// TIA Portal project "Projekt_Serhii_Bodnia" (V19)
// Vorlageprojekt für das Buch mit Zielsystem S7-1200

(* hardware
DEVICE "S7-1200-Station_1"  S7-1200 Station
   slot 0: "Baugruppenträger_0"  Rack  V1.0
   slot 1: "PLC_1"  CPU 1211C DC/DC/DC  6ES7 211-1AE40-0XB0  V4.1
DEVICE "HMI_1"  KTP900 Basic PN
   slot 0: "HMI_1"  KTP900 Basic PN  6AV2 123-2JB03-0AX0  17.0.0.0
   slot 1: "HMI_RT_1"  KTP900 Basic PN  6AV2 123-2JB03-0AX0  17.0.0.0
   slot 5: "HMI_1.IE_CP_1"  PROFINET Interface  17.0.0.0
      slot 1: "PROFINET Schnittstelle_1"  PROFINET Interface
         slot 1: "Port_1"  Port
*)

// ===== PLC "PLC_1"  CPU 1211C DC/DC/DC =====

VAR_GLOBAL   // PLC tag table "Standard-Variablentabelle"
   "System_Byte" AT %MB10 : Byte;
   "FirstScan" AT %M10.0 : Bool;
   "DiagStatusUpdate" AT %M10.1 : Bool;
   "Clock_Byte" AT %MB0 : Byte;
   "Clock_10Hz" AT %M0.0 : Bool;
   "Clock_5Hz" AT %M0.1 : Bool;
   "Clock_2.5Hz" AT %M0.2 : Bool;
   "Clock_2Hz" AT %M0.3 : Bool;
   "Clock_1.25Hz" AT %M0.4 : Bool;
   "Clock_1Hz" AT %M0.5 : Bool;
   "Clock_0.625Hz" AT %M0.6 : Bool;
   "Clock_0.5Hz" AT %M0.7 : Bool;
END_VAR

VAR_GLOBAL   // PLC tag table "Sensor"
   "Diffuse Sensor 0" AT %I0.0 : Bool;
   "Diffuse Sensor 1" AT %I0.1 : Bool;
   "Diffuse Sensor 2" AT %I0.2 : Bool;
   "Diffuse Sensor 3" AT %I0.3 : Bool;
   "Diffuse Sensor 4" AT %I0.4 : Bool;
   "Diffuse Sensor 5" AT %I0.5 : Bool;
   "Diffuse Sensor 6" AT %I0.6 : Bool;
   "Diffuse Sensor 7" AT %I0.7 : Bool;
   "Diffuse Sensor 8" AT %I1.0 : Bool;
   "Diffuse Sensor 9" AT %I1.1 : Bool;
   "Diffuse Sensor 10" AT %I1.2 : Bool;
   "Diffuse Sensor 11" AT %I1.3 : Bool;
   "Diffuse Sensor 12" AT %I1.4 : Bool;
   "Diffuse Sensor 13" AT %I1.5 : Bool;
   "Diffuse Sensor 14" AT %I1.6 : Bool;
   "Diffuse Sensor 15" AT %I1.7 : Bool;
   "Diffuse Sensor 16" AT %I2.0 : Bool;
   "Diffuse Sensor 17" AT %I2.1 : Bool;
   "Diffuse Sensor 18" AT %I2.2 : Bool;
   "Diffuse Sensor 19" AT %I2.3 : Bool;
   "Diffuse Sensor 20" AT %I2.4 : Bool;
   "Diffuse Sensor 21" AT %I2.5 : Bool;
   "Diffuse Sensor 22" AT %I2.6 : Bool;
   "Diffuse Sensor 23" AT %I2.7 : Bool;
   "Diffuse Sensor 24" AT %I3.0 : Bool;
   "Diffuse Sensor 25" AT %I3.1 : Bool;
   "Diffuse Sensor 26" AT %I3.2 : Bool;
   "Diffuse Sensor 27" AT %I3.3 : Bool;
   "Diffuse Sensor 29" AT %I3.4 : Bool;
   "Emergency Stop 0" AT %I3.6 : Bool;
   "Emergency Stop 1" AT %I3.7 : Bool;
   "Emergency Stop 3" AT %I4.0 : Bool;
   "Left Positioner 1 (Clamped)" AT %I3.5 : Bool;
   "Pick & Place 0 (Box Detected)" AT %I4.1 : Bool;
   "Retroreflective Sensor 1" AT %I4.2 : Bool;
   "Retroreflective Sensor 5" AT %I4.4 : Bool;
   "Retroreflective Sensor 7" AT %I4.5 : Bool;
   "Retroreflective Sensor 10" AT %I4.6 : Bool;
   "Start Button 0" AT %I5.3 : Bool;
   "Start Button 1" AT %I5.0 : Bool;
   "Stop Button 0" AT %I5.1 : Bool;
   "Stop Button 1" AT %I5.2 : Bool;
   "Conveyor Scale 0 Weight (V)" AT %ID30 : Real;
   "Conveyor Scale 1 Weight (V)" AT %ID34 : Real;
   "Tank 1 (Flow Meter)" AT %ID38 : Real;
   "Tank 2 (Flow Meter)" AT %ID42 : Real;
   "Tank 1 (Level Meter)" AT %ID46 : Real;
   "Tank 2 (Level Meter)" AT %ID50 : Real;
   "Vision Sensor 1 (Value)" AT %ID54 : DInt;
   "Retroreflective Sensor 2" AT %I4.3 : Bool;
END_VAR

VAR_GLOBAL   // PLC tag table "Aktor"
   "Belt Conveyor (2m) 0" AT %Q0.0 : Bool;
   "Belt Conveyor (2m) 1" AT %Q0.1 : Bool;
   "Belt Conveyor (2m) 2" AT %Q0.2 : Bool;
   "Belt Conveyor (2m) 3" AT %Q0.3 : Bool;
   "Belt Conveyor (2m) 4" AT %Q0.4 : Bool;
   "Belt Conveyor (4m) 0" AT %Q0.7 : Bool;
   "Belt Conveyor (4m) 2" AT %Q1.0 : Bool;
   "Belt Conveyor (4m) 3" AT %Q1.1 : Bool;
   "Belt Conveyor (4m) 5" AT %Q1.2 : Bool;
   "Belt Conveyor (4m) 6" AT %Q1.3 : Bool;
   "Belt Conveyor (4m) 7" AT %Q1.4 : Bool;
   "Belt Conveyor (6m) 2" AT %Q1.5 : Bool;
   "Belt Conveyor (2m) 6" AT %Q0.5 : Bool;
   "Belt Conveyor (2m) 7" AT %Q0.6 : Bool;
   "Conveyor Scale 0 (+)" AT %Q1.6 : Bool;
   "Conveyor Scale 1 (+)" AT %Q1.7 : Bool;
   "Curved Belt Conveyor 1 CW" AT %Q2.0 : Bool;
   "Curved Belt Conveyor 0 CCW" AT %Q2.1 : Bool;
   "Left Positioner 1 (Clamp)" AT %Q2.2 : Bool;
   "Emitter 1 (Emit)" AT %Q2.3 : Bool;
   "Emitter 3 (Emit)" AT %Q2.4 : Bool;
   "Emitter 4 (Emit)" AT %Q2.5 : Bool;
   "Remover 0 (Remove)" AT %Q2.6 : Bool;
   "Remover 1 (Remove)" AT %Q2.7 : Bool;
   "Remover 2 (Remove)" AT %Q3.0 : Bool;
   "Remover 3 (Remove)" AT %Q3.1 : Bool;
   "Roller Conveyor (2m) 0" AT %Q3.2 : Bool;
   "Roller Conveyor (2m) 1" AT %Q3.3 : Bool;
   "Roller Conveyor (2m) 3" AT %Q3.4 : Bool;
   "Roller Conveyor (4m) 0" AT %Q3.5 : Bool;
   "Pusher 0" AT %Q3.6 : Bool;
   "Pusher 3" AT %Q3.7 : Bool;
   "Pivot Arm Sorter 0 Turn" AT %Q4.0 : Bool;
   "Pivot Arm Sorter 0 Belt (+)" AT %Q4.1 : Bool;
   "Pick & Place 0 (Grab)" AT %Q4.2 : Bool;
   "Start Button 0 (Light)" AT %Q4.3 : Bool;
   "Start Button 1 (Light)" AT %Q4.4 : Bool;
   "Stop Button 0 (Light)" AT %Q4.5 : Bool;
   "Stop Button 1 (Light)" AT %Q4.6 : Bool;
   "Stack Light 0 (Green)" AT %Q4.7 : Bool;
   "Stack Light 0 (Red)" AT %Q5.0 : Bool;
   "Stack Light 0 (Yellow)" AT %Q5.1 : Bool;
   "Stack Light 1 (Green)" AT %Q5.2 : Bool;
   "Stack Light 1 (Red)" AT %Q5.3 : Bool;
   "Stack Light 1 (Yellow)" AT %Q5.4 : Bool;
   "Warning Light 1" AT %Q5.5 : Bool;
   "Pick & Place 0  X Set Point (V)" AT %QD34 : Real;
   "Pick & Place 0  Y Set Point (V)" AT %QD30 : Real;
   "Pick & Place 0  Z Set Point (V)" AT %QD38 : Real;
   "Tank 1 (Fill Valve)" AT %QD46 : Real;
   "Tank 2 (Fill Valve)" AT %QD50 : Real;
   "Tank 1 (Discharge Valve)" AT %QD54 : Real;
   "Tank 2 (Discharge Valve)" AT %QD58 : Real;
END_VAR

VAR_GLOBAL   // PLC tag table "Merker"
   "FlOp_P_Activate" AT %I4.7 : Bool;
END_VAR

TYPE "Getränk"
   STRUCT
      Tankfüllvolumen : Real;
      Dosiervolumen : Real;
      VAR_Rezeptur : Int;
      VAR_Rezeptur_Datensatz : Int;
   END_STRUCT;
END_TYPE

DATA_BLOCK "FB_Laufzeit_DB"   // DB1
{ S7_Optimized_Access := 'TRUE' }
VERSION : 0.1
// stored: InstanceOfName FB_Laufzeit
"FB_Laufzeit"
BEGIN
END_DATA_BLOCK

DATA_BLOCK "FB_Transport_Band_DB_1"   // DB2
{ S7_Optimized_Access := 'TRUE' }
VERSION : 0.1
// stored: InstanceOfName FB_Transport_Band
"FB_Transport_Band"
BEGIN
END_DATA_BLOCK

DATA_BLOCK "GDB_PLC"   // DB3
{ S7_Optimized_Access := 'TRUE' }
VERSION : 0.1
   VAR
      Dosierung_Start_Linie_0 : Bool;
      Dosierung_Start_Linie_1 : Bool;
      Dosing_Activate_Linie_0 : Bool;
      Dosing_Activate_Linie_1 : Bool;
      Eingabe_Level_norm_Linie_0 : Real;
      Eingabe_Level_norm_Linie_1 : Real;
      Tank_0_Level_norm : Real;
      Tank_1_Level_norm : Real;
      Start_Modus_Hauptleitung : Bool;
      Start_Modus_Linie_0 : Bool;
      Licht_in_Betrieb : Bool;
      Licht_außer_Betrieb : Bool;
      Licht_Alarm : Bool;
      Start_Modus_Linie_1 : Bool;
      Stop_Modus_Hauptleitung : Bool;
      Stop_Modus_Linie_0 : Bool;
      Stop_Modus_Linie_1 : Bool;
      Not_Aus_Modus : Bool;
      Füllventil_closed_Linie_0 : Bool;
      Füllventil_closed_Linie_1 : Bool;
      Altuell_Gewicht_Linie_0 : Real;
      Altuell_Gewicht_Linie_1 : Real;
      Gesamtteile_Linie_0 : Int;
      Gesamtteile_Linie_1 : Int;
      Ausschuss_Linie_0 : Int;
      Ausschuss_Linie_1 : Int;
      Anzahl_Paletten : Int;
      Anzahl_Kanister_Packungbereich : Int;
      Anzahl_Kanister_Tr_Band_Halle_2 : Int;
      Tankfüllvolumen_0 : Real;
      Tankfüllvolumen_1 : Real;
      Dosiervolumen_0 : Real;
      Dosiervolumen_1 : Real;
      Ready_to_Send_Teil_Band_Linie_3_0 : Bool;
      Acknowledge_Teil_Greifen_Linie_0 : Bool;
      Palette_voll_Linie_0 : Bool;
      Palette_voll_Linie_1 : Bool;
      Ready_To_Receive_Teil_Palette_Linie_0 : Bool;
      Ready_To_Receive_Teil_Palette_Linie_1 : Bool;
      Ready_To_Send_Teil_Wage_Linie_0 : Bool;
      Ready_To_Send_Teil_Band_2_Linie_0 : Bool;
      Ready_to_Receive_Teil_Band_3_Linie_0 : Bool;
      Run_Hours : Int;
      Run_Minutes : Int;
      Run_Seconds : Int;
      Störung : Array[0..16] of Bool;
   END_VAR
BEGIN
END_DATA_BLOCK

DATA_BLOCK "FB_Tank_DB"   // DB4
{ S7_Optimized_Access := 'TRUE' }
VERSION : 0.1
// stored: InstanceOfName FB_Tank
"FB_Tank"
BEGIN
END_DATA_BLOCK

DATA_BLOCK "FB_Dose_Control_DB"   // DB5
{ S7_Optimized_Access := 'TRUE' }
VERSION : 0.1
// stored: InstanceOfName FB_Dose_Control
"FB_Dose_Control"
BEGIN
END_DATA_BLOCK

DATA_BLOCK "GDB_HMI"   // DB6
{ S7_Optimized_Access := 'TRUE' }
VERSION : 0.1
   VAR
      Meldung_HMI : Int;
      Quittierung_HMI : Int;
      Tankfüllvolumen_HMI : Int;
      Dosiervolumen_HMI : Int;
      Füllmenge_Linie_0 : Real;
      Füllmenge_Linie_1 : Real;
      Reset_Gesamtteile_0 : Bool;
      Reset_Gesamtteile_1 : Bool;
      Reset_Ausschluss_0 : Bool;
      Reset_Ausschluss_1 : Bool;
      NotAus_HMI : Bool;
      Haupt_Stop_HMI : Bool;
   END_VAR
BEGIN
END_DATA_BLOCK

DATA_BLOCK "GDB_Getränk"   // DB7
{ S7_Optimized_Access := 'TRUE' }
VERSION : 0.1
   VAR
      Getränk_Linie_0 : "Getränk";
      Getränk_Linie_1 : "Getränk";
   END_VAR
BEGIN
END_DATA_BLOCK

DATA_BLOCK "FB_Transport_Band_DB_2"   // DB8
{ S7_Optimized_Access := 'TRUE' }
VERSION : 0.1
// stored: InstanceOfName FB_Transport_Band
"FB_Transport_Band"
BEGIN
END_DATA_BLOCK

DATA_BLOCK "FB_Mode_Manager_DB"   // DB9
{ S7_Optimized_Access := 'TRUE' }
VERSION : 0.1
// stored: InstanceOfName FB_Mode_Manager
"FB_Mode_Manager"
BEGIN
END_DATA_BLOCK

DATA_BLOCK "FB_Transport_Band_DB"   // DB10
{ S7_Optimized_Access := 'TRUE' }
VERSION : 0.1
// stored: InstanceOfName FB_Transport_Band
"FB_Transport_Band"
BEGIN
END_DATA_BLOCK

DATA_BLOCK "FB_AbfüllmaschineBand_SCL_DB"   // DB11
{ S7_Optimized_Access := 'TRUE' }
VERSION : 0.1
// stored: InstanceOfName FB_AbfüllmaschineBand_SCL
"FB_AbfüllmaschineBand_SCL"
BEGIN
END_DATA_BLOCK

DATA_BLOCK "FB_Gewichtkontrolle_SCL_DB"   // DB12
{ S7_Optimized_Access := 'TRUE' }
VERSION : 0.1
// stored: InstanceOfName FB_Gewichtkontrolle_SCL
"FB_Gewichtkontrolle_SCL"
BEGIN
END_DATA_BLOCK

DATA_BLOCK "FB_Transport_Band_DB_3"   // DB13
{ S7_Optimized_Access := 'TRUE' }
VERSION : 0.1
// stored: InstanceOfName FB_Transport_Band
"FB_Transport_Band"
BEGIN
END_DATA_BLOCK

DATA_BLOCK "FB_Sortierabschnitt_DB"   // DB14
{ S7_Optimized_Access := 'TRUE' }
VERSION : 0.1
// stored: InstanceOfName FB_Sortierabschnitt
"FB_Sortierabschnitt"
BEGIN
END_DATA_BLOCK

DATA_BLOCK "FB_Transport_Band_DB_4"   // DB15
{ S7_Optimized_Access := 'TRUE' }
VERSION : 0.1
// stored: InstanceOfName FB_Transport_Band
"FB_Transport_Band"
BEGIN
END_DATA_BLOCK

DATA_BLOCK "FB_Band mit Positionierleisten_DB"   // DB16
{ S7_Optimized_Access := 'TRUE' }
VERSION : 0.1
// stored: InstanceOfName FB_Band mit Positionierleisten
"FB_Band mit Positionierleisten"
BEGIN
END_DATA_BLOCK

DATA_BLOCK "FB_Palette_Linie_0_DB"   // DB17
{ S7_Optimized_Access := 'TRUE' }
VERSION : 0.1
// stored: InstanceOfName FB_Palette_Linie
"FB_Palette_Linie"
BEGIN
END_DATA_BLOCK

DATA_BLOCK "FB_Pick & Place_DB"   // DB18
{ S7_Optimized_Access := 'TRUE' }
VERSION : 0.1
// stored: InstanceOfName FB_Pick & Place
"FB_Pick & Place"
BEGIN
END_DATA_BLOCK

DATA_BLOCK "FB_Tank_DB_1"   // DB19
{ S7_Optimized_Access := 'TRUE' }
VERSION : 0.1
// stored: InstanceOfName FB_Tank
"FB_Tank"
BEGIN
END_DATA_BLOCK

DATA_BLOCK "FB_AbfüllmaschineBand_SCL_DB_1"   // DB20
{ S7_Optimized_Access := 'TRUE' }
VERSION : 0.1
// stored: InstanceOfName FB_AbfüllmaschineBand_SCL
"FB_AbfüllmaschineBand_SCL"
BEGIN
END_DATA_BLOCK

DATA_BLOCK "FB_Dose_Control_DB_1"   // DB21
{ S7_Optimized_Access := 'TRUE' }
VERSION : 0.1
// stored: InstanceOfName FB_Dose_Control
"FB_Dose_Control"
BEGIN
END_DATA_BLOCK

DATA_BLOCK "FB_Gewichtkontrolle_SCL_DB_1"   // DB22
{ S7_Optimized_Access := 'TRUE' }
VERSION : 0.1
// stored: InstanceOfName FB_Gewichtkontrolle_SCL
"FB_Gewichtkontrolle_SCL"
BEGIN
END_DATA_BLOCK

DATA_BLOCK "FB_Transport_Band_DB_5"   // DB23
{ S7_Optimized_Access := 'TRUE' }
VERSION : 0.1
// stored: InstanceOfName FB_Transport_Band
"FB_Transport_Band"
BEGIN
END_DATA_BLOCK

DATA_BLOCK "FB_Transport_Band_DB_6"   // DB24
{ S7_Optimized_Access := 'TRUE' }
VERSION : 0.1
// stored: InstanceOfName FB_Transport_Band
"FB_Transport_Band"
BEGIN
END_DATA_BLOCK

DATA_BLOCK "FB_Transport_Band_DB_7"   // DB25
{ S7_Optimized_Access := 'TRUE' }
VERSION : 0.1
// stored: InstanceOfName FB_Transport_Band
"FB_Transport_Band"
BEGIN
END_DATA_BLOCK

DATA_BLOCK "FB_Transportbad mit Verzögerung_DB"   // DB26
{ S7_Optimized_Access := 'TRUE' }
VERSION : 0.1
// stored: InstanceOfName FB_Transportbad mit Verzögerung
"FB_Transportbad mit Verzögerung"
BEGIN
END_DATA_BLOCK

DATA_BLOCK "FB_Transport_T-Band_DB"   // DB27
{ S7_Optimized_Access := 'TRUE' }
VERSION : 0.1
// stored: InstanceOfName FB_Transport_T-Band
"FB_Transport_T-Band"
BEGIN
END_DATA_BLOCK

DATA_BLOCK "FB_Transportbad mit Verzögerung_DB_1"   // DB28
{ S7_Optimized_Access := 'TRUE' }
VERSION : 0.1
// stored: InstanceOfName FB_Transportbad mit Verzögerung
"FB_Transportbad mit Verzögerung"
BEGIN
END_DATA_BLOCK

FUNCTION_BLOCK "FB_Gewichtkontrolle_SCL"   // FB1, SCL
{ S7_Optimized_Access := 'TRUE' }
VERSION : 0.1
   VAR_INPUT
      Start_Mode : Bool;
      Stop_Mode : Bool;
      NotAus_Mode : Bool;
      LS_Einlauf : Bool;
      LS_Mitte : Bool;
      LS_Auslauf : Bool;
      LS_Wage : Bool;
      LS_Pusher : Bool;
      Gewichtsskala : Real;
      Referenz_Gewicht : Real;
      Reset_CTU_Gesamtteile : Bool;
      Reset_CTU_Ausschuss : Bool;
      Quittierung : Bool;
   END_VAR
   VAR_OUTPUT
      Wage_Band : Bool;
      Pusher_Band : Bool;
      Gewicht_Kg : Real;
      Remoover : Bool;
      Pusher : Bool;
      Out_Gesamtteile : Int;
      Out_Ausschuss : Int;
      Ready_To_Send_Teil : Bool;
      Störung : Bool;
   END_VAR
   VAR
      iSchritt : Int;
      Trigger_Pos_LS_Einlauf : R_TRIG;
      Trigger_Neg_LS_Auslauf : F_TRIG;
      Trigger_Pos_LS_Mitte : R_TRIG;
      Trigger_Neg_LS_Mitte : F_TRIG;
      Trigger_Neg_LS_Wage : F_TRIG;
      Trigger_Neg_LS_Pusher : F_TRIG;
      TON_weit_Wiegung_1000ms : TON_TIME;
      TON_Puscher_100ms : TON_TIME;
      TON_Ende_weit_1000ms : TON_TIME;
      TOF_2000ms : TOF_TIME;
      Actuell_Gewicht : Real;
      Gewicht_Norm : Real;
      Speichen_Gewicht : Real;
      Gesamtteile : Int;
      Ausschuss : Int;
      TON_Störung_LS_Wage : TON_TIME;
      TON_Störung_LS_Mitte : TON_TIME;
      TON_Störung_LS_Pusher : TON_TIME;
      TON_Störung_Auslauf : TON_TIME;
      M_Störung : Bool;
      M_Wage_Band : Bool;
      M_Pusher_Band : Bool;
   END_VAR
   VAR CONSTANT
      Toleranz : Real := 1.02;
   END_VAR
BEGIN
   REGION NotAus & Störung
       IF #NotAus_Mode OR #M_Störung THEN
           // Bei Not-Aus or Störung sofortiger Rücksprung in den Initialschritt (Schritt 0)
           #iSchritt := 0;
       END_IF;
   END_REGION

   REGION Reset
       IF #Reset_CTU_Gesamtteile OR #NotAus_Mode OR "FirstScan" THEN
           // Gesamtteilezähler zurücksetzen: bei HMI-Anforderung, Not-Aus oder Erstaufruf
           #Gesamtteile := 0;
       END_IF;

       IF #Reset_CTU_Ausschuss OR #NotAus_Mode OR "FirstScan" THEN
           // Ausschusszähler zurücksetzen: bei HMI-Anforderung, Not-Aus oder Erstaufruf
           #Ausschuss := 0;

       END_IF;

   END_REGION

   REGION Flankenabfragen
       #Trigger_Pos_LS_Einlauf(CLK := #LS_Einlauf); 
       #Trigger_Pos_LS_Mitte(CLK := #LS_Mitte);     
       #Trigger_Neg_LS_Mitte(CLK := #LS_Mitte);
       #Trigger_Neg_LS_Auslauf(CLK := #LS_Auslauf);
       #Trigger_Neg_LS_Wage(CLK := #LS_Wage);
       #Trigger_Neg_LS_Pusher(CLK := #LS_Pusher);
   END_REGION

   REGION Timers
       // Wiegezeit: 500ms Wartezeit für stabile Gewichtsmessung (Schritt 2)
       #TON_weit_Wiegung_1000ms(IN := (#iSchritt = 2),
                                PT := T#500ms);
       // Pusher-Impuls: 100ms Aktivierungszeit für Pusher-Zylinder (Schritt 11)
       #TON_Puscher_100ms(IN := #iSchritt = 11,
                          PT := T#100ms);
       // Remover-Wartezeit: 1000ms bis Remover das Ausschussteil aufgenommen hat (Schritt 12)
       #TON_Ende_weit_1000ms(IN := (#iSchritt = 12),
                             PT := T#1000ms);
       // Anzeigedauer Gewicht: Messwert 2 Sekunden nach Wiegung sichtbar halten (Schritt 2)
       #TOF_2000ms(IN := (#iSchritt = 2),
                   PT := T#2000ms);
       // Störungserkennung: wenn Licht_Sensors länger als 10s aktiv und Band läuft → Stau

       #TON_Störung_LS_Wage(IN := #LS_Wage AND #M_Wage_Band AND NOT #Stop_Mode,
                            PT := T#10s);
       #TON_Störung_LS_Mitte(IN := #LS_Mitte AND #M_Wage_Band AND NOT #Stop_Mode,
                             PT := T#10s);
       #TON_Störung_LS_Pusher(IN := #LS_Pusher AND #M_Pusher_Band AND NOT #Stop_Mode,
                             PT := T#10s);
       #TON_Störung_Auslauf(IN := #LS_Auslauf AND #M_Pusher_Band AND NOT #Stop_Mode,
                            PT := T#10s);

   END_REGION

   REGION Scalierung_Gewicht
       // Rohwert Wiegezelle (0–10 V analog) auf 0–20 kg normieren und skalieren
       #Gewicht_Norm := NORM_X(MIN := 0.0, VALUE := #Gewichtsskala, MAX := 10.0);
       #Actuell_Gewicht:= SCALE_X_REAL(MIN := 0.0, VALUE := #Gewicht_Norm, MAX := 20.0);

   END_REGION

   REGION Meldungen
       // Störungserkennung: wenn LS_Einlauf oder LS_Auslauf länger als 10s aktiv und Band läuft → Stau
       IF (#TON_Störung_LS_Wage.Q OR #TON_Störung_LS_Mitte.Q)
           OR (#TON_Störung_LS_Pusher.Q OR #TON_Störung_Auslauf.Q) THEN
           // Störungsmerker setzen
           #M_Störung := TRUE;
       END_IF;
       // Störung über HMI quittieren: Bit des Quittierungswortes (HMI_Quittierung.%X0)
       IF #Quittierung THEN
           #M_Störung := FALSE;
       END_IF;

   END_REGION


   REGION Schrittkette
       CASE #iSchritt OF
           0:  // Initialschritt: Warten auf Teil am Einlauf UND Startmodus
               IF #Trigger_Pos_LS_Einlauf.Q AND #Start_Mode THEN
                   #iSchritt := 1;
               END_IF;
           1:  // Waageband läuft; Gesamtteilezähler erhöhen, wenn Teil die Waage erreicht
               IF #Trigger_Neg_LS_Wage.Q THEN
                   #Gesamtteile := #Gesamtteile + 1;
                   #iSchritt := 2;
               END_IF;
           2:  // Wiegung: Band gestoppt, 500ms warten für stabile Messwerterfassung
               IF #TON_weit_Wiegung_1000ms.Q THEN
                   #Speichen_Gewicht := #Actuell_Gewicht;
                   #iSchritt := 3;
               END_IF;
           3:  // Gewichtsprüfung: bei LS_Mitte-Flanke Toleranzband prüfen
               // Toleranzband: Referenz/1,02 ≤ Gewicht ≤ Referenz*1,02 (±2%)
               IF #Trigger_Pos_LS_Mitte.Q THEN
                   IF (#Speichen_Gewicht <= #Referenz_Gewicht * #Toleranz)
                       AND (#Speichen_Gewicht >= #Referenz_Gewicht / #Toleranz) THEN
                       #iSchritt := 4;
                   ELSE
                       #Ausschuss := #Ausschuss + 1;
                       #iSchritt := 10;
                   END_IF;
               END_IF;
           4:  // Waageband UND Pusherband laufen; warten bis Teil Mitte verlässt
               IF #Trigger_Neg_LS_Mitte.Q THEN
                   #iSchritt := 5;
               END_IF;
           5: // Waageband AUS, Pusherband läuft; Teil zum Auslauf befördern
              // Sobald Teil den Auslauf verlässt: prüfen ob schon nächstes Teil wartet
               IF #Trigger_Neg_LS_Auslauf.Q THEN
                   IF #LS_Einlauf THEN
                       #iSchritt := 1; // Nächstes Teil sofort verarbeiten
                   ELSE
                       #iSchritt := 0; // Kein weiteres Teil → Initialschritt
                   END_IF;
               END_IF;
           10: // Ausschleuspfad: Pusherband läuft; Teil zum Pusher-Lichtschranke befördern
               IF #Trigger_Neg_LS_Pusher.Q THEN
                   #iSchritt := 11;
               END_IF;
           11: // Pusher aktivieren für 100ms (Ausschussteil seitwärts ausschieben)
               IF #TON_Puscher_100ms.Q THEN
                   #iSchritt := 12;
               END_IF;
           12: // Remover aktiv für 1000ms (Ausschussteil endgültig entfernen)
               IF #TON_Ende_weit_1000ms.Q THEN
                   #iSchritt := 0; // Zurück zum Initialschritt
               END_IF;

       END_CASE;

   END_REGION
   REGION Actoren
       // 1. Wage_Band
       #M_Wage_Band := (#iSchritt = 1 OR #iSchritt = 3 OR #iSchritt = 4 OR #iSchritt = 10) AND NOT #Stop_Mode;
       #Wage_Band := #M_Wage_Band;
       // 2. Pusher_Band
       #M_Pusher_Band:= (#iSchritt = 4 OR #iSchritt = 5 OR #iSchritt = 10 OR #iSchritt =11 OR #iSchritt =12) AND NOT #Stop_Mode;
       #Pusher_Band := #M_Pusher_Band;
       // 3. Pusher
       #Pusher := #iSchritt = 11;
       // 4. Remover
       #Remoover := #iSchritt = 12;
       // 5. Zähler
       #Out_Gesamtteile := #Gesamtteile;
       #Out_Ausschuss := #Ausschuss;
       // 
       #Ready_To_Send_Teil := NOT #Stop_Mode AND (#iSchritt = 4 OR  #iSchritt = 5);

   END_REGION
   REGION Gewicht anzeige
       // Gewichtsanzeige: Messwert 2 Sekunden nach Wiegung anzeigen, danach auf 0 setzen
       // TOF bleibt 2s aktiv nachdem Schritt 2 verlassen wurde
       IF #TOF_2000ms.Q THEN
           #Gewicht_Kg := #Speichen_Gewicht;
       ELSE
           #Gewicht_Kg := 0.0;
       END_IF;
   END_REGION
END_FUNCTION_BLOCK

FUNCTION_BLOCK "FB_Tank"   // FB2, FBD
TITLE = FB_Tank
{ S7_Optimized_Access := 'TRUE' }
VERSION : 0.1
// Füllstand einstellen per HMI
   VAR_INPUT
      "Tank (Levelmeter)" : Real;
      Input_HMI_Level : Real;
      HMI_acknowledge : Int;
      Start_Mode : Bool;
      Not_Aus : Bool;
      Stop_Mode : Bool;
   END_VAR
   VAR_OUTPUT
      "Tank (Füllventil)" : Real;
      Füllventil_closed : Bool;
      HMI_Meldung : Int;
   END_VAR
   VAR
      Input_Level : Real;
      Diff_Level : Real;
      valve_value : Real;
      intermediate_result : Real;
      dynamic_value : Real;
      IEC_TON_message : TON_TIME;
      SR_message_level_reached : Bool;
      SR_message_valve_open : Bool;
      complete_open : Bool;
      complete_closed : Bool;
      dynamic_open : Bool;
      SR_acknowledge : Bool;
   END_VAR
   VAR_TEMP   // added for the SCL form of the ladder/FBD networks
      _w1 : Bool;
   END_VAR
BEGIN

REGION Network 1: Input level / Acknowledgement
   // Der Sollwert wird nur geschrieben, wenn der Tank leer ist, oder der Füllstand in der HMI quittiert wurde.
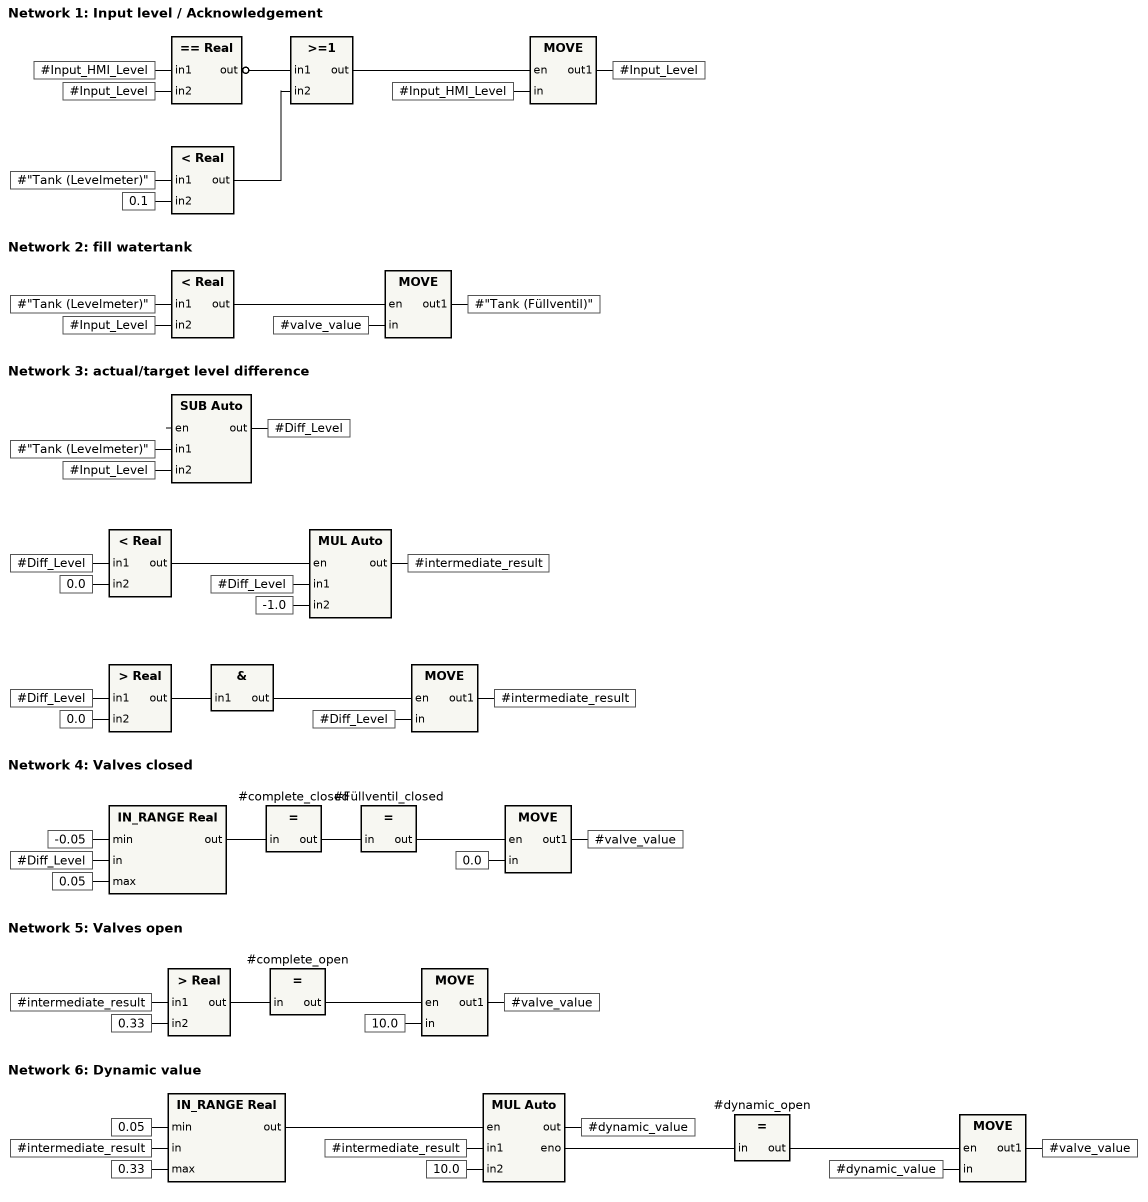
   IF NOT (#Input_HMI_Level = #Input_Level) OR (#"Tank (Levelmeter)" < 0.1) THEN
       #Input_Level := #Input_HMI_Level;
   END_IF;
END_REGION

REGION Network 2: fill watertank
   // Füllen, solange Ist-Wert kleiner Soll-Wert
   IF #"Tank (Levelmeter)" < #Input_Level THEN #"Tank (Füllventil)" := #valve_value; END_IF;
END_REGION

REGION Network 3: actual/target level difference
   // Erfassen der Differenz zwischen Soll und Ist, ein negatives Ergebnis wird invertiert
   #Diff_Level := #"Tank (Levelmeter)" - #Input_Level;
   IF #Diff_Level < 0.0 THEN #intermediate_result := #Diff_Level * (-1.0); END_IF;
   IF #Diff_Level > 0.0 THEN #intermediate_result := #Diff_Level; END_IF;
END_REGION

REGION Network 4: Valves closed
   // Ist die Differenz kleiner als 0.05, ist der Valve Value 0.0 (komplett geschlossen)
   #complete_closed := (-0.05 <= #Diff_Level) AND (#Diff_Level <= 0.05);
   #Füllventil_closed := #complete_closed;
   IF #complete_closed THEN #valve_value := 0.0; END_IF;
END_REGION

REGION Network 5: Valves open
   // Ist die Differenz größer als 0.33, ist der valve value 10.0 (komplett offen)
   #complete_open := #intermediate_result > 0.33;
   IF #complete_open THEN #valve_value := 10.0; END_IF;
END_REGION

REGION Network 6: Dynamic value
   // dynamischer Valve Value ab 0.33 Differenz  bis 0.05 Differenz mit Verstärkung 10
   #_w1 := (0.05 <= #intermediate_result) AND (#intermediate_result <= 0.33);
   IF #_w1 THEN #dynamic_value := #intermediate_result * 10.0; END_IF;
   #dynamic_open := #_w1;
   IF #_w1 THEN #valve_value := #dynamic_value; END_IF;
END_REGION

REGION Network 7 (SCL): Not Aus, Stop und Tank-Überfüllscnutz
   //Not Aus und Stop 
   IF #Not_Aus THEN
       #Füllventil_closed := TRUE;
       #"Tank (Füllventil)" := 0.0;
       #valve_value := 0.0;
       #dynamic_value := 0.0;
       #dynamic_open := FALSE;
   ELSIF #Stop_Mode THEN
       #valve_value := 0.0;
       #"Tank (Füllventil)" := 0.0;
       #Füllventil_closed := TRUE;
   END_IF;

   // Tank-Überfüllscnutz
   IF #"Tank (Levelmeter)" >= 0.98 THEN
       #valve_value := 0.0;
       #"Tank (Füllventil)" := 0.0;
       #Füllventil_closed := TRUE;
   END_IF;
END_REGION
END_FUNCTION_BLOCK

FUNCTION_BLOCK "FB_Dose_Control"   // FB3, SCL
{ S7_Optimized_Access := 'TRUE' }
VERSION : 0.1
   VAR_INPUT
      Trigger_Start : Bool;
      Flow_Raw : Real;
      Target_Volume : Real;
      Not_Aus : Bool;
   END_VAR
   VAR_OUTPUT
      Discharge_Valve : Real;
      Dosing_Status : Bool;
      Füllmenge : Real;
   END_VAR
   VAR
      sTrigger : R_TRIG;
      Accumulated_Vol : Real;
      Dosing_Activate : Bool;
      Stat_Timer_Reset : TOF_TIME;
   END_VAR
   VAR CONSTANT
      C_Q_MAX_M3_S : Real := 0.3543;   // Maximaler Volumenstrom (10V = 0,3543 m³/s) [m³/s]
      C_OB30_ZEIT_S : Real := 0.01;   // OB30-Zykluszeit (muss mit CPU-Konfig. übereinstimmen) [s]
      C_M3_TO_L : Real := 1000.0;   // Umrechnungsfaktor Kubikmeter → Liter [l/m³]
      C_U_MAX_V : Real := 10.0;   // Analogbereich Maximum [V]
   END_VAR
BEGIN
   REGION Flankenabfragen
       // Steigende Flanke des Dosierstarts erfassen (Trigger_Start ist ein Impuls)
       #sTrigger(CLK := #Trigger_Start);
   END_REGION

   REGION Timers
       // TOF: nach Ende der Dosierung bleibt .Q für 1 Sekunde TRUE
       // → verhindert sofortiges Rücksetzen von Accumulated_Vol nach Dosierungsende 
       #Stat_Timer_Reset(IN := #Dosing_Activate,
                         PT := T#1s);

   END_REGION

   REGION #Not_Aus
       IF #Not_Aus THEN
           #Accumulated_Vol := 0.0;
           #Dosing_Activate := FALSE;
       END_IF;


   END_REGION

   REGION Dosierung
       // Dosierung starten: nur bei steigender Flanke UND wenn Dosierung noch nicht läuft
       IF #sTrigger.Q AND NOT #Dosing_Activate THEN
           #Accumulated_Vol := 0.0;
           #Dosing_Activate := TRUE;
       END_IF;
       IF #Dosing_Activate THEN
           // Volumenstrom integrieren über die OB30-Zykluszeit
           // Formel: ΔVol = Flow_Raw / 10.0 * 0.3543 * 0.01 * 1000

           #Accumulated_Vol := #Accumulated_Vol + (#Flow_Raw / #C_U_MAX_V * #C_Q_MAX_M3_S * #C_OB30_ZEIT_S * #C_M3_TO_L);
           IF #Accumulated_Vol < (#Target_Volume * 0.85) THEN
               // Zweistufige Ventilsteuerung: Großhub bis 85% des Zielvolumens, dann Kleinhub
               // Schnellfüllung: Ventil weit offen
               #Discharge_Valve := 2.0;
           ELSE
               // Feindosierung: Ventil fast geschlossen
               #Discharge_Valve := 0.05;
           END_IF;
           IF #Accumulated_Vol >= (#Target_Volume - 0.2) THEN
               // Dosierung beenden, wenn Zielvolumen (mit 0,2l Vorhalt) erreicht
               #Dosing_Activate := FALSE;
           END_IF;
       ELSE
           // Keine aktive Dosierung: Ventil vollständig schließen
           #Discharge_Valve := 0.0;
       END_IF;

       IF NOT #Dosing_Activate AND NOT #Stat_Timer_Reset.Q THEN
           // Volumenrücksetzung: 1 Sekunde nach Dosierungsende (TOF-Fenster)
           // Verhindert sofortiges Löschen der Anzeige nach Abfüllung
           #Accumulated_Vol := 0.0;
       END_IF;

   END_REGION


   // Statusausgaben für HMI-Anzeige
   #Dosing_Status := #Dosing_Activate; // TRUE während aktiver Dosierung
   #Füllmenge := #Accumulated_Vol; // Aktuell abgefüllte Menge für HMI
END_FUNCTION_BLOCK

FUNCTION_BLOCK "FB_Transportbad mit Verzögerung"   // FB4, SCL
{ S7_Optimized_Access := 'TRUE' }
VERSION : 0.1
   VAR_INPUT
      LS_Einlauf : Bool;
      LS_Auslauf : Bool;
      Start_Modus : Bool;
      Stop_Modus : Bool;
      NotAus_Modus : Bool;
      Nächste_Band_belegt : Bool;
      Quittierung : Bool;
   END_VAR
   VAR_OUTPUT
      Band : Bool;
      Ready_to_Send_Teil : Bool;
      Störung : Bool;
   END_VAR
   VAR
      FlOp_Pos_LS_Einlauf : R_TRIG;
      FlOp_Neg_LS_Auslauf : F_TRIG;
      FlOp_Pos_LS_Auslauf : R_TRIG;
      Teil_auf_Band : Int;
      M_Band : Bool;
      M_Störung : Bool;
      M_Teil_wartet : Bool;
      TON_Störung_LS_Einlauf : TON_TIME;
      TON_Störung_LS_Ausauf : TON_TIME;
   END_VAR
BEGIN
   REGION Flankenabfragen
       // Flankenauswertungen für Einlauf- und Auslaufsensoren
       #FlOp_Pos_LS_Einlauf(CLK := #LS_Einlauf);
       #FlOp_Neg_LS_Auslauf(CLK := #LS_Auslauf);
       #FlOp_Pos_LS_Auslauf(CLK := #LS_Auslauf);

   END_REGION

   REGION Timers
       // Störungserkennung: wenn LS_Einlauf oder LS_Auslauf länger als 10s aktiv und Band läuft → Stau
       #TON_Störung_LS_Einlauf(IN := #LS_Einlauf AND #M_Band AND NOT #Stop_Modus,
                               PT := T#10s);
       #TON_Störung_LS_Ausauf(IN := #LS_Auslauf AND #M_Band AND NOT #Stop_Modus,
                              PT := T#10s);
   END_REGION

   REGION Meldungen
       // Störungserkennung: wenn LS_Einlauf oder LS_Auslauf länger als 3s aktiv und Band läuft → Stau
       IF (#Teil_auf_Band > 3 OR #TON_Störung_LS_Einlauf.Q OR #TON_Störung_LS_Ausauf.Q) AND NOT #M_Teil_wartet THEN
           // Störungsmerker setzen
           #M_Störung := TRUE;
       END_IF;
       // Störung über HMI quittieren: Bit des Quittierungswortes (HMI_Quittierung)
       IF #Quittierung THEN
           #M_Störung := FALSE;
       END_IF;

   END_REGION

   REGION Erfassung der Anzahl der Teileauf dem Band
       // Teilezähler: Inkrementierung bei jedem neuen Teil von beiden Einläufen
       IF #Start_Modus AND NOT #Stop_Modus AND #FlOp_Pos_LS_Einlauf.Q THEN
           #Teil_auf_Band := #Teil_auf_Band + 1;
       END_IF;
       // Dekrementierung wenn Teil den Auslauf verlässt
       IF #Start_Modus AND NOT #Stop_Modus AND #FlOp_Neg_LS_Auslauf.Q AND #Teil_auf_Band > 0 THEN
           #Teil_auf_Band := #Teil_auf_Band - 1;
       END_IF;
       // Not-Aus: Teilezähler zurücksetzen
       IF #NotAus_Modus THEN
           #Teil_auf_Band := 0;
       END_IF;
   END_REGION

   REGION Band
       // Wartelogik: Teil am Auslauf detektiert UND nächstes Band ist belegt → warten
       // M_Teil_wartet ist kombinatorisch (kein Halteglied), reagiert sofort auf Statusänderung

       IF #Start_Modus AND #LS_Auslauf AND #Nächste_Band_belegt THEN
           // Teil muss warten: nächstes Band noch besetzt
           #M_Teil_wartet := TRUE;
       ELSE
           // Nächstes Band frei: kann weiterfahren
           #M_Teil_wartet := FALSE;
       END_IF;
       // Bandsteuerung: läuft wenn Teile auf Band oder neues Teil angekommen
       IF #Start_Modus AND (#FlOp_Pos_LS_Einlauf.Q OR #Teil_auf_Band > 0) THEN
           #M_Band := True;
       ELSE
           #M_Band := FALSE;
       END_IF;
       IF #NotAus_Modus OR #M_Störung THEN
           #M_Band := FALSE;
       END_IF;

   END_REGION

   REGION Ready_To_Send & Ready_To_Receive
       // Weitergabesignal: Teil wartet am Auslauf auf freies nächstes Band
       // Dieses Signal wird vom nachgelagerten Band (FB_Transportbad) ausgewertet

       #"Ready_to_Send_Teil" := #M_Teil_wartet;

   END_REGION

   REGION Aktoren
       // Physischer Ausgang:  Band stoppt bei: Stopp-Modus ODER Teil wartet auf nächstes Band
       // Automatischer Wiederanlauf wenn Nächste_Band_belegt FALSE wird
       #Band := #M_Band AND NOT #M_Teil_wartet AND NOT #Stop_Modus;
       #Störung := #M_Störung;

   END_REGION
END_FUNCTION_BLOCK

FUNCTION_BLOCK "FB_Transport_Band"   // FB5, SCL
{ S7_Optimized_Access := 'TRUE' }
VERSION : 0.1
   VAR_INPUT
      LS_Einlauf : Bool;
      LS_Ausauf : Bool;
      Start_Modus : Bool;
      Stop_Modus : Bool;
      NotAus_Modus : Bool;
      Quittierung : Bool;
   END_VAR
   VAR_OUTPUT
      Band : Bool;
      Störung : Bool;
   END_VAR
   VAR
      FlOp_Pos_LS_Einlauf : R_TRIG;
      FlOp_Neg_LS_Auslauf : F_TRIG;
      FlOp_Pos_LS_Auslauf : R_TRIG;
      Teil_auf_Band : Int;
      M_Band : Bool;
      TON_Störung_Einlauf : TON_TIME;
      TON_Störung_Auslauf : TON_TIME;
      M_Störung : Bool;
   END_VAR
BEGIN

   REGION Flankenabfragen
       // Alle Flanken müssen am Anfang des Bausteins aktualisiert werden
       #FlOp_Pos_LS_Einlauf(CLK := #LS_Einlauf);
       #FlOp_Neg_LS_Auslauf(CLK := #LS_Ausauf);
       #FlOp_Pos_LS_Auslauf(CLK := #LS_Ausauf);

   END_REGION

   REGION Timers
       // Störungserkennung: wenn LS_Auslauf länger als 10s aktiv und Band läuft → Stau
       #TON_Störung_Auslauf(IN := #LS_Ausauf AND #M_Band AND NOT #Stop_Modus,
                            PT := T#10s);
       #TON_Störung_Einlauf(IN := #LS_Einlauf AND #M_Band AND NOT #Stop_Modus,
                            PT := T#10s);
   END_REGION

   REGION Meldungen
       // Störungserkennung: wenn LS_Einlauf oder LS_Auslauf länger als 10s aktiv und Band läuft → Stau
       IF  (#Teil_auf_Band > 3 OR #TON_Störung_Auslauf.Q OR #TON_Störung_Einlauf.Q)  THEN
           // Störungsmerker setzen
           #M_Störung := TRUE;
       END_IF;
       // Störung über HMI quittieren: Bit des Quittierungswortes (HMI_Quittierung)
       IF #Quittierung THEN
           #M_Störung := FALSE;
       END_IF;

   END_REGION

   REGION Erfassung der Anzahl der Teileauf dem Band
       // Teil kommt auf Band: steigende Flanke am Einlauf (nur im aktiven Betrieb)
       IF #Start_Modus AND #FlOp_Pos_LS_Einlauf.Q THEN
           #Teil_auf_Band := #Teil_auf_Band + 1;
       END_IF;
       // Teil verlässt Band: fallende Flanke am Auslauf (Zähler nie unter 0)
       IF #Start_Modus AND #FlOp_Neg_LS_Auslauf.Q AND #Teil_auf_Band > 0 THEN
           #Teil_auf_Band := #Teil_auf_Band - 1;
       END_IF;
       // Not-Aus: Teilezähler sofort zurücksetzen
       IF #NotAus_Modus OR #M_Störung THEN
           #Teil_auf_Band := 0;
       END_IF;
   END_REGION

   REGION Band
       // Band einschalten: wenn Startmodus UND (neues Teil oder Teile noch auf Band)
       IF #Start_Modus AND (#FlOp_Pos_LS_Einlauf.Q OR #Teil_auf_Band > 0) THEN
           #M_Band := True;
       ELSE
           // Kein Teil auf Band: Band abschalten
           #M_Band := FALSE;
       END_IF;
       // Not-Aus und Störung: Band sofort abschalten
       IF #NotAus_Modus OR #M_Störung THEN
           #M_Band := FALSE;
       END_IF;

   END_REGION

   REGION Aktoren
       // Physischer Ausgang: Band läuft nur wenn Merker gesetzt UND kein Stopp-Modus
       #Band := #M_Band AND NOT #Stop_Modus;
       #Störung := #M_Störung;
   END_REGION
END_FUNCTION_BLOCK

FUNCTION_BLOCK "FB_Sortierabschnitt"   // FB6, SCL
{ S7_Optimized_Access := 'TRUE' }
VERSION : 0.1
   VAR_INPUT
      LS_Einlauf_Band_0 : Bool;
      LS_Auslauf_Band_0 : Bool;
      LS_Einlauf_Band_1 : Bool;
      LS_Auslauf_Band_1 : Bool;
      LS_Vision_Sensor : Bool;
      LS_Arm_0 : Bool;
      Vision_Sensor : DInt;
      Produktart_Linie_0 : Int;
      Produktart_Linie_1 : Int;
      Start_Modus : Bool;
      Stop_Modus : Bool;
      Not_Aus_Modus : Bool;
      Quittierung : Bool;
   END_VAR
   VAR_OUTPUT
      Band_0 : Bool;
      Band_1 : Bool;
      Arm_turn_0 : Bool;
      Arm_Band_0 : Bool;
      Remover : Bool;
      Anzahl_Kanister : Int;
      Störung : Bool;
   END_VAR
   VAR
      Buffer : Array[0..5] of DInt;
      Count : Int;
      Current_Art : DInt;
      Rezeptur_Art_0 : DInt;
      Rezeptur_Art_1 : DInt;
      i : Int;
      FlOp_Pos_LS_Vision_Sensor : R_TRIG;
      FlOp_Pos_LS_Arm_0 : R_TRIG;
      FlOp_Neg_LS_Einlauf_Band_0 : F_TRIG;
      FlOp_Pos_LS_Einlauf_Band_1 : R_TRIG;
      FlOp_Neg_LS_Auslauf_Band_1 : F_TRIG;
      "FlOp_Neg_LS_Auslauf_Band_0 (1)" : F_TRIG;
      "FlOp_Neg_LS_Auslauf_Band_0 (2)" : F_TRIG;
      TP_Remover : TP_TIME;
      TON_Störung_LS_Einlauf_Band_0 : TON_TIME;
      TON_Störung_LS_Auslauf_Band_0 : TON_TIME;
      TON_Störung_LS_Einlauf_Band_1 : TON_TIME;
      TON_Störung_LS_Auslauf_Band_1 : TON_TIME;
      TON_Störung_LS_Vision_Sensor : TON_TIME;
      TON_Störung_LS_Arm_0 : TON_TIME;
      Teil_auf_Band_0 : Int;
      Teil_auf_Band_1 : Int;
      M_Band_0 : Bool;
      M_Band_1 : Bool;
      M_Arm_turn_0 : Bool;
      M_Arm_Band_0 : Bool;
      CTU_Kanister : CTU_INT;
      M_Störung : Bool;
   END_VAR
BEGIN
   REGION Flankenabfragen
       // Flankenauswertungen für alle Sensoren des Sortierabschnitts
       #FlOp_Neg_LS_Einlauf_Band_0(CLK := #"LS_Einlauf_Band_0");
       #"FlOp_Neg_LS_Auslauf_Band_0 (1)"(CLK := #LS_Auslauf_Band_0 );
       #"FlOp_Neg_LS_Auslauf_Band_0 (2)"(CLK := #LS_Einlauf_Band_1 );
       #FlOp_Pos_LS_Einlauf_Band_1(CLK := #LS_Einlauf_Band_1);
       #FlOp_Neg_LS_Auslauf_Band_1(CLK := #LS_Auslauf_Band_1);
       #FlOp_Pos_LS_Vision_Sensor(CLK := #LS_Vision_Sensor);
       #FlOp_Pos_LS_Arm_0(CLK := #LS_Arm_0);

   END_REGION

   REGION Zähler
       // Fertigteile zählen: Inkrementierung bei jeder Fallende-Flanke am Auslauf Band 1
       #CTU_Kanister(CU:= #FlOp_Neg_LS_Auslauf_Band_1.Q,
                     R:= "FirstScan" OR #Not_Aus_Modus,
                     PV:=0);
                  END_REGION